(* CODESYS project TA5450_AB_2_2_2.project

Project tree, tasks and I/O mapping:
  PLC_AC500_V3 : PM5630-2ETH, ABB Automation Products GmbH, order no. 1SAP131000R0278, version 3.2.2.0
    application Application
      libraries: Util, * (System)
      task Task (cyclic, interval t#10ms, priority 15, watchdog t#20ms x 1) calls PLC_PRG
      task VISU_TASK (cyclic, interval 100 ms, priority 16) calls VisuElems.Visu_Prg
      CheckConfigurationObject
      program PLC_PRG [ST]
      program LD_example [LD]
      program FBD_example [FBD]
      program CFC_example [CFC]
      global variables GVL
      visualisation Visualization
      image pool ImagePool
      Symbols
    IO_Bus : I/O-Bus, ABB Automation Products GmbH, version 3.2.1.0
      DA501 : DA501, ABB Automation Products GmbH, order no. 1SAPx50700R0001, version 3.2.1.0
          input  xDI_08_DA501 : BOOL  // Digital inputs DI8 - DI15.Digital input DI8
          input  xDI_09_DA501 : BOOL  // Digital inputs DI8 - DI15.Digital input DI9
          input  xDI_10_DA501 : BOOL  // Digital inputs DI8 - DI15.Digital input DI10
          input  xDI_11_DA501 : BOOL  // Digital inputs DI8 - DI15.Digital input DI11
          input  xAI_00_DA501 : INT  // Analog input AI0+
          input  xAI_01_DA501 : INT  // Analog input AI1+
          output xDO_16_DA501 : BOOL  // Digital outputs DC16 - DC23.Digital output DC16
          output xDO_17_DA501 : BOOL  // Digital outputs DC16 - DC23.Digital output DC17
          output xDO_18_DA501 : BOOL  // Digital outputs DC16 - DC23.Digital output DC18
          output xDO_19_DA501 : BOOL  // Digital outputs DC16 - DC23.Digital output DC19
          output xDO_21_DA501 : BOOL  // Digital outputs DC16 - DC23.Digital output DC21
          output xDO_22_DA501 : BOOL  // Digital outputs DC16 - DC23.Digital output DC22
          output xDO_23_DA501 : BOOL  // Digital outputs DC16 - DC23.Digital output DC23
          unmapped channels: Input0, Input1, Input2, Output0, Output1, Digital inputs DI0 - DI15, Analog input AI0+, Analog input AI1+, Analog input AI2+, Analog input AI3+, Digital inputs DC16 - DC23, Reserved, Analog output AO0+, Analog output AO1+, Reserved, Digital outputs DC16 - DC23, Reserved, Digital inputs DI0 - DI7, Digital inputs DI8 - DI15, Digital inputs DC16 - DC23, Reserved, Analog input AI2+, Analog input AI3+, Fast counter input, Digital outputs DC16 - DC23, Reserved, Analog output AO0+, Analog output AO1+, Reserved, Fast counter output, Digital inputs DI0 - DI7, Digital inputs DI8 - DI15, Digital inputs DC16 - DC23, Analog input AI0+, Analog input AI1+, Analog input AI2+, Analog input AI3+, Digital outputs DC16 - DC23, Analog output AO0+, Analog output AO1+,
            Reserved
    Interfaces : Interfaces, ABB Automation Products GmbH, version 3.2.0.0
      COM_1 : COM 1, ABB Automation Products GmbH, version 3.2.0.0
        CAA_SerialCom : CAA SerialCom, ABB Automation Products GmbH, version 3.2.0.0
      CAN
      Ethernet : Ethernet, ABB Automation Products GmbH, version 3.2.0.0
        ETH1 : IP Settings, ABB Automation Products GmbH, version 3.2.0.0
          NetConfig : NetConfig, ABB Automation Products GmbH, version 3.2.0.0
        ETH2 : IP Settings, ABB Automation Products GmbH, version 3.2.0.0
          NetConfig_1 : NetConfig, ABB Automation Products GmbH, version 3.2.0.0
        Protocols : Client Protocols, ABB Automation Products GmbH, version 3.2.0.0
    Extension_Bus : Extension Bus, ABB Automation Products GmbH, version 3.2.0.0
      CM579_PNIO : CM579-PNIO, ABB Automation Products GmbH, order no. 1SAPx70901R0101, version 3.2.0.0
          settings: Slot number = 1
        PNIO_Controller : PROFINET-IO-Controller, ABB Automation Products GmbH, version 3.2.0.0
            settings: IP address = [192, 168, 0, 1]; Subnet Mask = [255, 255, 255, 0]; Gateway Address = [0, 0, 0, 0]; First IP Address = [192, 168, 0, 2]; Last IP Address = [192, 168, 0, 254]; Default Subnet Mask = [255, 255, 255, 0]; Default Gateway Address = [0, 0, 0, 0]; PackageSizeDesc.Number of devices = 1; PackageSizeDesc.Max. number of API = 1; PackageSizeDesc.Max. number of modules = 2; PackageSizeDesc.Max. number of submodules = 1; PackageSizeDesc.Max. number of RecData = 59; OrderID = '1SAPx70901R0101'
          CI502_PNIO_Device : CI502-PNIO-Device, ABB Automation Products GmbH, order no. 1SAPx20700R0001, version 3.2.0.0
              settings: Slave parameters.Identification.IP address = [192,168,0,2]; Slave parameters.Identification.Subnet mask = [255,255,255,0]; Slave parameters.Identification.Default gateway = [0,0,0,0]; Slave parameters.Identification.MAC address = [16#00,16#00,16#00,16#00,16#00,16#00]; Slave parameters.Identification.Station name = 'ci502-pn-02'; Slave parameters.Watchdog interval = 3; PDPortDataCheck.PeerStationName = ''; PDPortDataCheck.PeerStationName = ''; CRParameters.aCRPrm.Input_FrameLength = 18; CRParameters.aCRPrm.Input_IODataSize = 12; CRParameters.aCRPrm.Input_PSDataSize = 5; CRParameters.aCRPrm.Input_CSDataSize = 5; CRParameters.aCRPrm.Input_ulProp = 2; CRParameters.aCRPrm.Input_SendClockFact = 32; CRParameters.aCRPrm.Input_ReductionRatio = 4; CRParameters.aCRPrm.Output_FrameLength = 26; CRParameters.aCRPrm.Output_IODataSize = 20; CRParameters.aCRPrm.Output_PSDataSize = 1; CRParameters.aCRPrm.Output_CSDataSize = 1; CRParameters.aCRPrm.Output_ulProp = 2; CRParameters.aCRPrm.Output_SendClockFact = 32; CRParameters.aCRPrm.Output_ReductionRatio = 4; ARUUID = [72,189,233,212,83,232,168,78,179,79,33,17,12,11,1,46]; FSParamUuidData = [65,233,148,249,66,213,79,77,141,40,157,119,47,114,151,59]; SubModuleIoDesc_CI502 DIM1.SubModuleIoDesc.Input_IOPSSize = 1; SubModuleIoDesc_CI502 DIM1.SubModuleIoDesc.Input_IOCSSize = 1; SubModuleIoDesc_CI502 DIM1.SubModuleIoDesc.Output_Type = 0; SubModuleIoDesc_CI502 DIM1.SubModuleIoDesc.Output_IOCRRef = 1; SubModuleIoDesc_CI502 DIM1.SubModuleIoDesc.Output_IOCRRefOppositeDirecction = 0; SubModuleIoDesc_ci502-pn-00.SubModuleIoDesc.Input_IOPSSize = 1; SubModuleIoDesc_ci502-pn-00.SubModuleIoDesc.Input_IOCSSize = 1; SubModuleIoDesc_ci502-pn-00.SubModuleIoDesc.Input_FrameOffset = 1; SubModuleIoDesc_ci502-pn-00.SubModuleIoDesc.Input_CSOffset = 1; SubModuleIoDesc_ci502-pn-00.SubModuleIoDesc.Output_Type = 0; SubModuleIoDesc_ci502-pn-00.SubModuleIoDesc.Output_IOCRRef = 1; SubModuleIoDesc_ci502-pn-00.SubModuleIoDesc.Output_IOCRRefOppositeDirecction = 0; SubModuleIoDesc_port-001.SubModuleIoDesc.Input_IOPSSize = 1; SubModuleIoDesc_port-001.SubModuleIoDesc.Input_IOCSSize = 1; SubModuleIoDesc_port-001.SubModuleIoDesc.Input_FrameOffset = 2; SubModuleIoDesc_port-001.SubModuleIoDesc.Input_CSOffset = 2;
                SubModuleIoDesc_port-001.SubModuleIoDesc.Output_Type = 0; SubModuleIoDesc_port-001.SubModuleIoDesc.Output_IOCRRef = 1; SubModuleIoDesc_port-001.SubModuleIoDesc.Output_IOCRRefOppositeDirecction = 0; SubModuleIoDesc_port-002.SubModuleIoDesc.Input_IOPSSize = 1; SubModuleIoDesc_port-002.SubModuleIoDesc.Input_IOCSSize = 1; SubModuleIoDesc_port-002.SubModuleIoDesc.Input_FrameOffset = 3; SubModuleIoDesc_port-002.SubModuleIoDesc.Input_CSOffset = 3; SubModuleIoDesc_port-002.SubModuleIoDesc.Output_Type = 0; SubModuleIoDesc_port-002.SubModuleIoDesc.Output_IOCRRef = 1; SubModuleIoDesc_port-002.SubModuleIoDesc.Output_IOCRRefOppositeDirecction = 0
            CI502_IO : CI502-IO, ABB Automation Products GmbH, order no. 1SAPx20700R0001, version 3.2.0.0
                settings: Module parameters.Slot number = 1; swapInfoInputs = [10,2,12,2,10,2]; swapInfoOutputs = [10,2,12,4,10,2]; 8-bit digital input_DPRAM = [0, 0, 0, 0, 192, 0, 0, 0, 10, 0, 8, 0]; 8-bit digital input_DPRAM = [8, 0, 0, 0, 200, 0, 0, 0, 10, 0, 8, 0]; Fast Counter: Actual value 1_DPRAM = [16, 0, 0, 0, 224, 0, 0, 0, 12, 0, 32, 0]; Fast Counter: Actual value 2_DPRAM = [48, 0, 0, 0, 0, 1, 0, 0, 12, 0, 32, 0]; Fast Counter: State byte 1_DPRAM = [80, 0, 0, 0, 32, 1, 0, 0, 10, 0, 8, 0]; Fast Counter: State byte 2_DPRAM = [88, 0, 0, 0, 40, 1, 0, 0, 10, 0, 8, 0]; 8-bit digital output_DPRAM = [0, 0, 0, 0, 224, 0, 0, 0, 10, 0, 8, 0]; 8-bit digital output_DPRAM = [8, 0, 0, 0, 232, 0, 0, 0, 10, 0, 8, 0]; Fast Counter: Start value 1_DPRAM = [16, 0, 0, 0, 0, 1, 0, 0, 12, 0, 32, 0]; Fast Counter: End value 1_DPRAM = [48, 0, 0, 0, 32, 1, 0, 0, 12, 0, 32, 0]; Fast Counter: Start value 2_DPRAM = [80, 0, 0, 0, 64, 1, 0, 0, 12, 0, 32, 0]; Fast Counter: End value 2_DPRAM = [112, 0, 0, 0, 96, 1, 0, 0, 12, 0, 32, 0]; Fast Counter: Control byte 1_DPRAM = [144, 0, 0, 0, 128, 1, 0, 0, 10, 0, 8, 0]; Fast Counter: Control byte 2_DPRAM = [152, 0, 0, 0, 136, 1, 0, 0, 10, 0, 8, 0]; SubModuleIoDesc_CI502 Input/Output.SubModuleIoDesc.Input_IODataSize = 12; SubModuleIoDesc_CI502 Input/Output.SubModuleIoDesc.Input_IOPSSize = 1; SubModuleIoDesc_CI502 Input/Output.SubModuleIoDesc.Input_IOCSSize = 1; SubModuleIoDesc_CI502 Input/Output.SubModuleIoDesc.Input_FrameOffset = 4; SubModuleIoDesc_CI502 Input/Output.SubModuleIoDesc.Input_CSOffset = 4; SubModuleIoDesc_CI502 Input/Output.SubModuleIoDesc.Output_IOCRRef = 1; SubModuleIoDesc_CI502 Input/Output.SubModuleIoDesc.Output_IOCRRefOppositeDirecction = 0; SubModuleIoDesc_CI502 Input/Output.SubModuleIoDesc.Output_IODataSize = 20; SubModuleIoDesc_CI502 Input/Output.SubModuleIoDesc.Output_IOPSSize = 1; SubModuleIoDesc_CI502 Input/Output.SubModuleIoDesc.Output_IOCSSize = 1
                input  xDI_08_CI502 : BOOL  // 8-bit digital input.Channel 8
                input  xDI_09_CI502 : BOOL  // 8-bit digital input.Channel 9
                input  xDI_10_CI502 : BOOL  // 8-bit digital input.Channel 10
                input  xDI_11_CI502 : BOOL  // 8-bit digital input.Channel 11
                output xDO_08_CI502 : BOOL  // 8-bit digital output.Channel 8
                output xDO_09_CI502 : BOOL  // 8-bit digital output.Channel 9
                output xDO_10_CI502 : BOOL  // 8-bit digital output.Channel 10
                output xDO_11_CI502 : BOOL  // 8-bit digital output.Channel 11
                output xDO_13_CI502 : BOOL  // 8-bit digital output.Channel 13
                output xDO_14_CI502 : BOOL  // 8-bit digital output.Channel 14
                output xDO_15_CI502 : BOOL  // 8-bit digital output.Channel 15
                unmapped channels: 8-bit digital input, 8-bit digital input, Fast Counter: Actual value 1, Fast Counter: Actual value 2, Fast Counter: State byte 1, Fast Counter: State byte 2, 8-bit digital output, 8-bit digital output, Fast Counter: Start value 1, Fast Counter: End value 1, Fast Counter: Start value 2, Fast Counter: End value 2, Fast Counter: Control byte 1, Fast Counter: Control byte 2
      Slot 2
  Panel_CP600 : CP600 Control Panel, ABB Automation Products GmbH, order no. 1SAP500900R0001, version 2.8.0.0
    CP6607_project_and_HMI_demo
  text list GlobalTextList
  5ce3da45-db07-42e7-a21c-a00fff4ed8f6|C:\Users\DEU214980\Desktop\Folders\Projekte\Training Case V3\V3_Project\bmp\3ADR333332V0015_DA501.png
  5ce3da45-db07-42e7-a21c-a00fff4ed8f6|C:\Users\DEU214980\Desktop\Folders\Projekte\Training Case V3\V3_Project\bmp\3ADR333220V0015_CI502-PNIO.png
*)

// PLC_AC500_V3/Application/GVL
{attribute 'qualified_only'}
VAR_GLOBAL
	Pot_AI1: INT;
	Pot_AI2: INT;
END_VAR

// PLC_AC500_V3/Application/PLC_PRG
PROGRAM PLC_PRG
VAR
END_VAR

LD_example();
FBD_example();
CFC_example();

END_PROGRAM

// PLC_AC500_V3/Application/LD_example
PROGRAM LD_example
VAR
(* Function Block Instances *)
	TON2: TON;	(* Timer On Delay *)
	CTU2: CTU;	(* Counter Up *)

(* FB outputs *)
	tTimer_Value2: TIME;(* Elapsed Time *)
	wCounter_Value2: WORD;(* Current Counter Value *)
	xCTU2_LimitReached: BOOL;
END_VAR

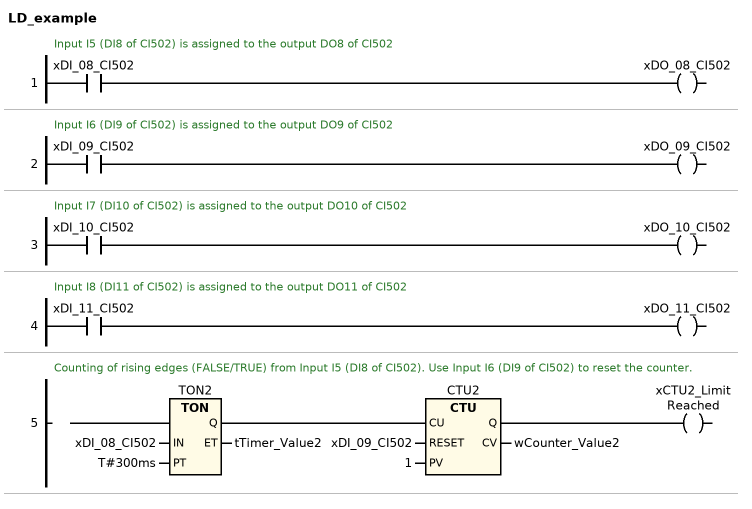
// NETWORK 1
// Input I5 (DI8 of CI502) is assigned to the output DO8 of CI502
xDO_08_CI502 := xDI_08_CI502;

// NETWORK 2
// Input I6 (DI9 of CI502) is assigned to the output DO9 of CI502
xDO_09_CI502 := xDI_09_CI502;

// NETWORK 3
// Input I7 (DI10 of CI502) is assigned to the output DO10 of CI502
xDO_10_CI502 := xDI_10_CI502;

// NETWORK 4
// Input I8 (DI11 of CI502) is assigned to the output DO11 of CI502
xDO_11_CI502 := xDI_11_CI502;

// NETWORK 5
// Counting of rising edges (FALSE/TRUE) from Input I5 (DI8 of CI502). Use Input I6 (DI9 of CI502) to reset the counter.
TON2(IN := xDI_08_CI502, PT := T#300ms, ET => tTimer_Value2); // TON
CTU2(CU := TON2.Q, RESET := xDI_09_CI502, PV := 1, CV => wCounter_Value2); // CTU
xCTU2_LimitReached := CTU2.Q;

END_PROGRAM

// PLC_AC500_V3/Application/FBD_example
PROGRAM FBD_example
VAR

(* Function Block Instances *)
	TON1: TON;	(* Timer On Delay *)
	CTU1: CTU;	(* Counter Up *)

(* FB outputs *)
	tTimer_Value1: TIME;(* Elapsed Time *)
	wCounter_Value1: WORD;(* Current Counter Value *)
	xCTU1_LimitReached: BOOL;
END_VAR

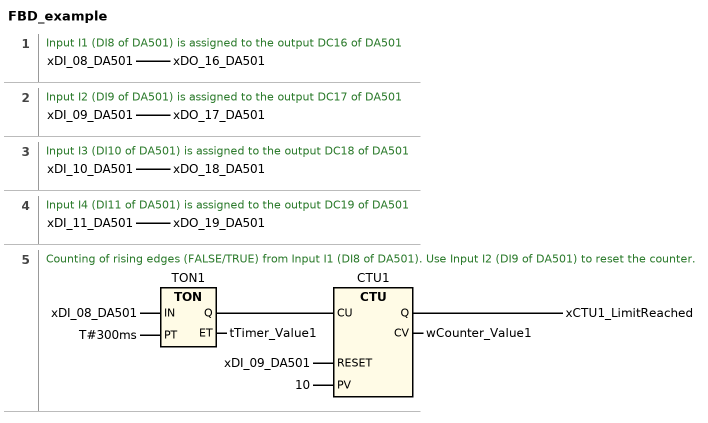
// NETWORK 1
// Input I1 (DI8 of DA501) is assigned to the output DC16 of DA501
xDO_16_DA501 := xDI_08_DA501;

// NETWORK 2
// Input I2 (DI9 of DA501) is assigned to the output DC17 of DA501
xDO_17_DA501 := xDI_09_DA501;

// NETWORK 3
// Input I3 (DI10 of DA501) is assigned to the output DC18 of DA501
xDO_18_DA501 := xDI_10_DA501;

// NETWORK 4
// Input I4 (DI11 of DA501) is assigned to the output DC19 of DA501
xDO_19_DA501 := xDI_11_DA501;

// NETWORK 5
// Counting of rising edges (FALSE/TRUE) from Input I1 (DI8 of DA501). Use Input I2 (DI9 of DA501) to reset the counter.
TON1(IN := xDI_08_DA501, PT := T#300ms, ET => tTimer_Value1); // TON
CTU1(CU := TON1.Q, RESET := xDI_09_DA501, PV := 10, CV => wCounter_Value1); // CTU
xCTU1_LimitReached := CTU1.Q;

END_PROGRAM

// PLC_AC500_V3/Application/CFC_example
PROGRAM CFC_example
VAR
(* Function Block Instances *)
	LIMITALARM1: LIMITALARM;
	LIMITALARM2: LIMITALARM;

END_VAR
VAR // added by the converter: edge detectors and wires of the graphical bodies
    _w1, _w2 : ANY;
END_VAR

// Scaling and  generation of limit alarms for AI2 signal  (AI1 analog input of DA501). The signal ranges (overflow, underflow, normal) are indicated by outputs DCO13 - DO15 of  CI502)
_w1 := LIMIT(xAI_01_DA501, 0, 27000) / 2700;
GVL.Pot_AI2 := _w1;
LIMITALARM2(IN := _w1, HIGH := 8, LOW := 2); // LIMITALARM
xDO_13_CI502 := LIMITALARM2.O;
xDO_15_CI502 := LIMITALARM2.U;
// Scaling and  generation of limit alarms for AI1 signal  (AI0 analog input of DA501). The signal ranges (overflow, underflow, normal) are indicated by outputs DC21 - DC23 of  DA501)
_w2 := LIMIT(xAI_00_DA501, 0, 27000) / 2700;
LIMITALARM1(IN := _w2, HIGH := 8, LOW := 2); // LIMITALARM
xDO_14_CI502 := LIMITALARM2.IL;
GVL.Pot_AI1 := _w2;
xDO_21_DA501 := LIMITALARM1.O;
xDO_23_DA501 := LIMITALARM1.U;
xDO_22_DA501 := LIMITALARM1.IL;

END_PROGRAM

// PLC_AC500_V3/Application/Visualization
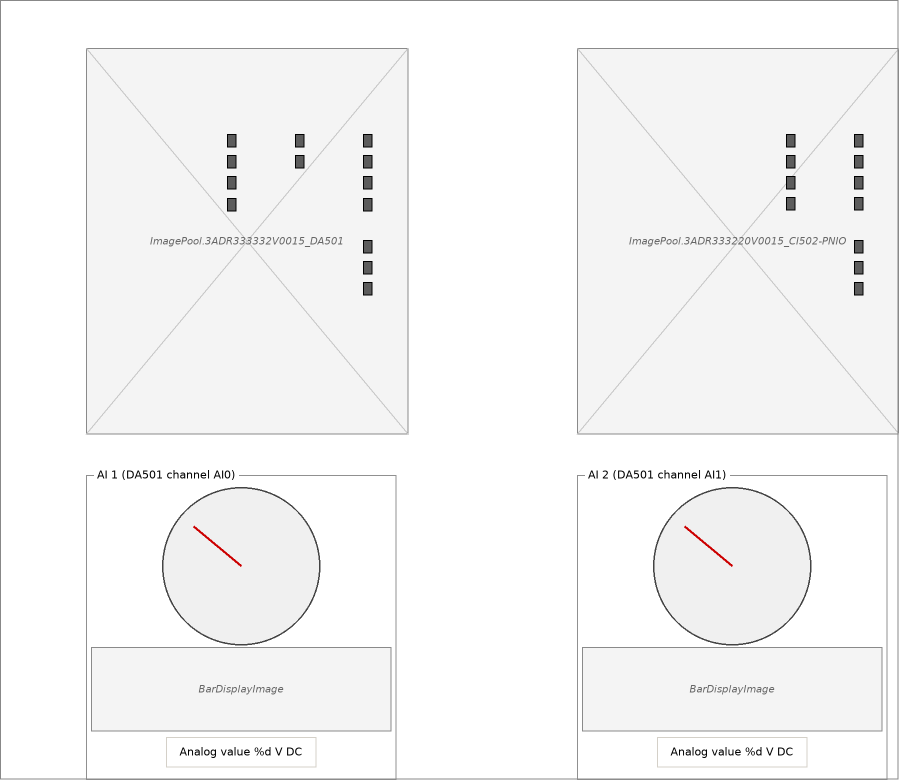
VISUALIZATION Visualization  // 899x780, background image VisuElems.IP_ElementImages.Rectangle
    GroupBox (86,467 310x313), "AI 1 (DA501 channel AI0)"
        Meter180 (5,20 300x158), value: GVL.Pot_AI1, style: Meter-Meter180-Gray, scale format: %.1f, scale 0..10
        BarDisplayImage (5,180 300x84), value: GVL.Pot_AI1, style: BarDisplayImage-Gray, scale format: %.1f, scale 0..10
        Textfield (80,270 150x30), "Analog value %d V DC", text variable: GVL.Pot_AI1
    GroupBox (577,467 310x313), "AI 2 (DA501 channel AI1)"
        Meter180 (5,20 300x158), value: GVL.Pot_AI2, style: Meter-Meter180-Gray, scale format: %.1f, scale 0..10
        BarDisplayImage (5,180 300x84), value: GVL.Pot_AI2, style: BarDisplayImage-Gray, scale format: %.1f, scale 0..10
        Textfield (80,270 150x30), "Analog value %d V DC", text variable: GVL.Pot_AI2
    Group (577,48 322x386)
        Image (0,0 322x386), image: ImagePool.3ADR333220V0015_CI502-PNIO
        RoundedRectangle (209,86 9x13), colour toggle: xDI_08_CI502
        RoundedRectangle (209,107 9x13), colour toggle: xDI_09_CI502
        RoundedRectangle (209,128 9x13), colour toggle: xDI_10_CI502
        RoundedRectangle (209,149 9x13), colour toggle: xDI_11_CI502
        RoundedRectangle (277,86 9x13), colour toggle: xDO_08_CI502
        RoundedRectangle (277,107 9x13), colour toggle: xDO_09_CI502
        RoundedRectangle (277,128 9x13), colour toggle: xDO_10_CI502
        RoundedRectangle (277,149 9x13), colour toggle: xDO_11_CI502
        RoundedRectangle (277,234 9x13), colour toggle: xDO_15_CI502
        RoundedRectangle (277,213 9x13), colour toggle: xDO_14_CI502
        RoundedRectangle (277,192 9x13), colour toggle: xDO_13_CI502
    Group (86,48 322x386)
        Image (0,0 322x386), image: ImagePool.3ADR333332V0015_DA501
        RoundedRectangle (141,86 9x13), colour toggle: xDI_08_DA501
        RoundedRectangle (141,107 9x13), colour toggle: xDI_09_DA501
        RoundedRectangle (141,128 9x13), colour toggle: xDI_10_DA501
        RoundedRectangle (141,150 9x13), colour toggle: xDI_11_DA501
        RoundedRectangle (277,86 9x13), colour toggle: xDO_16_DA501
        RoundedRectangle (277,107 9x13), colour toggle: xDO_17_DA501
        RoundedRectangle (277,128 9x13), colour toggle: xDO_18_DA501
        RoundedRectangle (277,150 9x13), colour toggle: xDO_19_DA501
        RoundedRectangle (277,192 9x13), colour toggle: xDO_21_DA501
        RoundedRectangle (277,213 9x13), colour toggle: xDO_22_DA501
        RoundedRectangle (277,234 9x13), colour toggle: xDO_23_DA501
        RoundedRectangle (209,86 9x13), colour toggle: xDO_21_DA501, invisible if: xDO_22_DA501 AND xDO_23_DA501
        RoundedRectangle (209,86 9x13), colour toggle: xDO_22_DA501, invisible if: xDO_21_DA501
        RoundedRectangle (209,107 9x13), colour toggle: xDO_13_CI502, invisible if: xDO_14_CI502 AND xDO_15_CI502
        RoundedRectangle (209,107 9x13), colour toggle: xDO_14_CI502, invisible if: xDO_13_CI502
END_VISUALIZATION
